(* Logix 5000 project; controller PLC_MCC1201_220AP1 vendor 1 type 14 code 164 rev 35.11; software revision 35.00; part 7 of 25 *)
(* tags used below, declared in another part *)
   B3 : DINT[102];
   HMI_Alarm_Reset : BOOL;   // HMI_Alarm_Reset
   HMI_MAN_CMD_WR : UDT_MAN_CMD_WR;
   LEHR_SPEED : ALIAS FOR N60[1];
   M210_M1_DR : AXIS_CIP_DRIVE;
   M211_M1_DR : AXIS_CIP_DRIVE;
   M212_M1_DR : AXIS_CIP_DRIVE;
   M213_M1_DR : AXIS_CIP_DRIVE;
   M2xx_CONVEYOR : MAC_CONVEYOR[20];
   M2xx_CONVEYOR_IN_MOTION : MAC_CONVEYOR_IN_MOTION[20];
   M2xx_CONVEYOR_OUT_MOTION : MAC_CONVEYOR_OUT_MOTION[20];
   TMP_dDirection : DINT;
   TMP_rAcc : REAL;
   TMP_rDec : REAL;
   TMP_rSpeed : REAL;
   TMP_xAlwaysOFF : BOOL;
   TMP_xRun : BOOL;
(* CommandLogic, continued *)

ROUTINE M210_Conveyor_Motion_Output   (* ladder *)
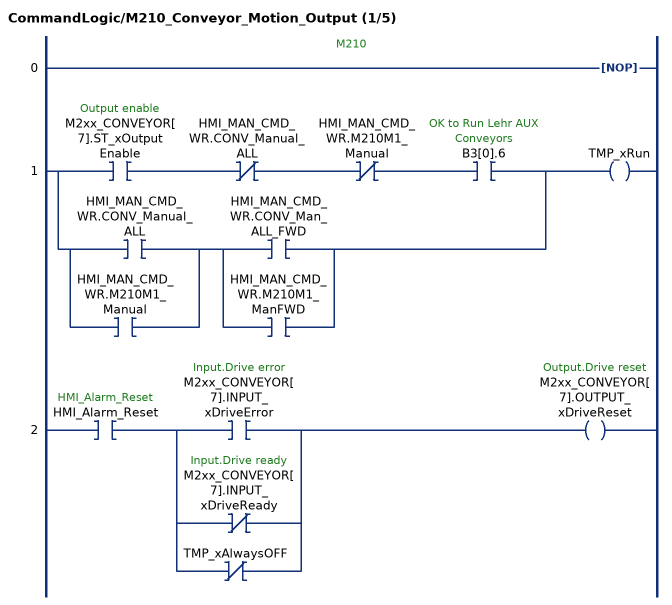
   // M210
   0: NOP();
   1: [XIC(M2xx_CONVEYOR[7].ST_xOutputEnable) XIO(HMI_MAN_CMD_WR.CONV_Manual_ALL) XIO(HMI_MAN_CMD_WR.M210M1_Manual) XIC(B3[0].6) ,[XIC(HMI_MAN_CMD_WR.CONV_Manual_ALL) ,XIC(HMI_MAN_CMD_WR.M210M1_Manual) ] [XIC(HMI_MAN_CMD_WR.CONV_Man_ALL_FWD) ,XIC(HMI_MAN_CMD_WR.M210M1_ManFWD) ] ]OTE(TMP_xRun);
   2: XIC(HMI_Alarm_Reset)[XIC(M2xx_CONVEYOR[7].INPUT_xDriveError) ,XIO(M2xx_CONVEYOR[7].INPUT_xDriveReady) ,XIO(TMP_xAlwaysOFF) ]OTE(M2xx_CONVEYOR[7].OUTPUT_xDriveReset);
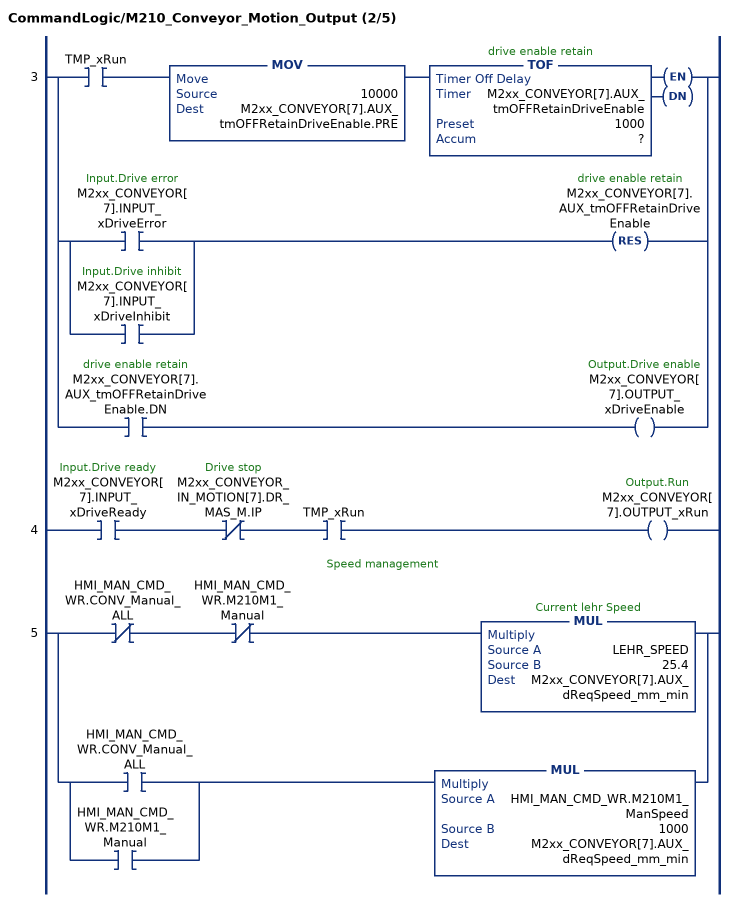
   3: [XIC(TMP_xRun) MOV(10000,M2xx_CONVEYOR[7].AUX_tmOFFRetainDriveEnable.PRE) TOF(M2xx_CONVEYOR[7].AUX_tmOFFRetainDriveEnable,?,?) ,[XIC(M2xx_CONVEYOR[7].INPUT_xDriveError) ,XIC(M2xx_CONVEYOR[7].INPUT_xDriveInhibit) ] RES(M2xx_CONVEYOR[7].AUX_tmOFFRetainDriveEnable) ,XIC(M2xx_CONVEYOR[7].AUX_tmOFFRetainDriveEnable.DN) OTE(M2xx_CONVEYOR[7].OUTPUT_xDriveEnable) ];
   4: XIC(M2xx_CONVEYOR[7].INPUT_xDriveReady)XIO(M2xx_CONVEYOR_IN_MOTION[7].DR_MAS_M.IP)XIC(TMP_xRun)OTE(M2xx_CONVEYOR[7].OUTPUT_xRun);
   // Speed management
   5: [XIO(HMI_MAN_CMD_WR.CONV_Manual_ALL) XIO(HMI_MAN_CMD_WR.M210M1_Manual) MUL(LEHR_SPEED,25.4,M2xx_CONVEYOR[7].AUX_dReqSpeed_mm_min) ,[XIC(HMI_MAN_CMD_WR.CONV_Manual_ALL) ,XIC(HMI_MAN_CMD_WR.M210M1_Manual) ] MUL(HMI_MAN_CMD_WR.M210M1_ManSpeed,1000,M2xx_CONVEYOR[7].AUX_dReqSpeed_mm_min) ];
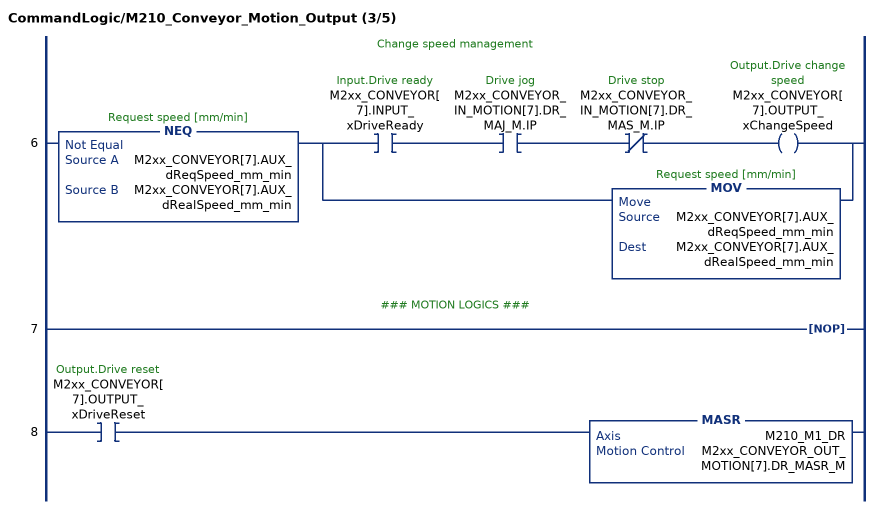
   // Change speed management
   6: NEQ(M2xx_CONVEYOR[7].AUX_dReqSpeed_mm_min,M2xx_CONVEYOR[7].AUX_dRealSpeed_mm_min)[XIC(M2xx_CONVEYOR[7].INPUT_xDriveReady) XIC(M2xx_CONVEYOR_IN_MOTION[7].DR_MAJ_M.IP) XIO(M2xx_CONVEYOR_IN_MOTION[7].DR_MAS_M.IP) OTE(M2xx_CONVEYOR[7].OUTPUT_xChangeSpeed) ,MOV(M2xx_CONVEYOR[7].AUX_dReqSpeed_mm_min,M2xx_CONVEYOR[7].AUX_dRealSpeed_mm_min) ];
   // ### MOTION LOGICS ###
   7: NOP();
   8: XIC(M2xx_CONVEYOR[7].OUTPUT_xDriveReset)MASR(M210_M1_DR,M2xx_CONVEYOR_OUT_MOTION[7].DR_MASR_M);
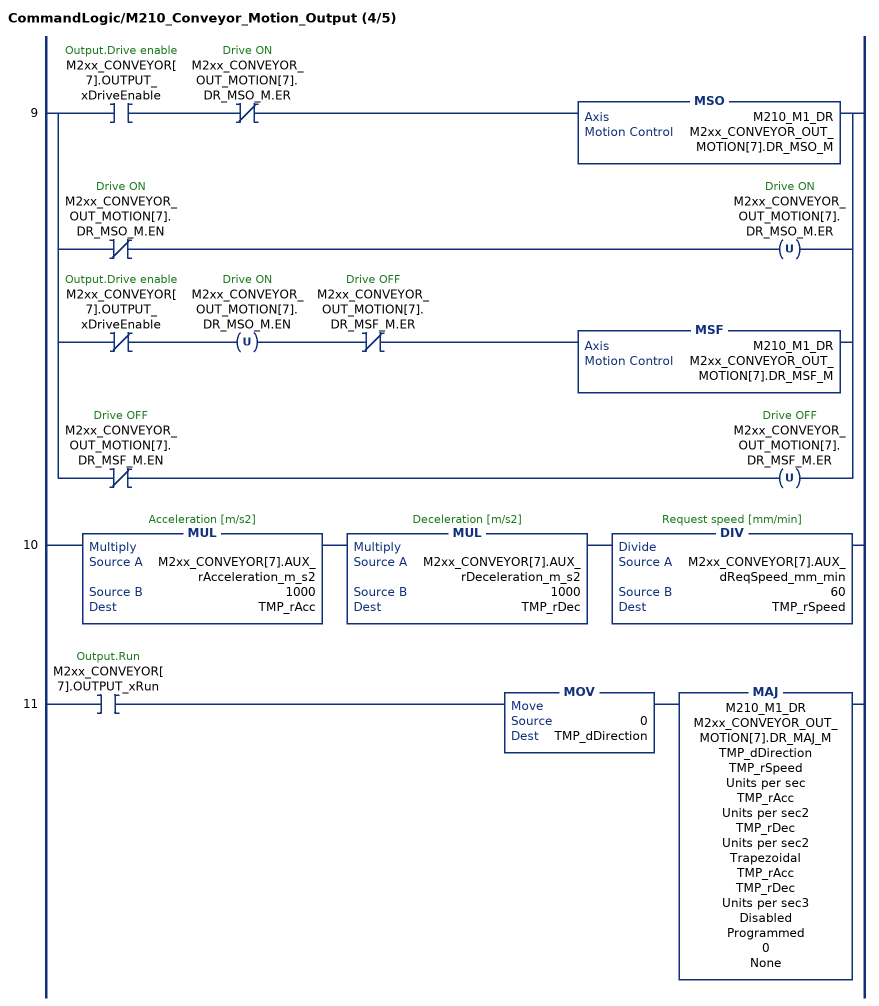
   9: [XIC(M2xx_CONVEYOR[7].OUTPUT_xDriveEnable) XIO(M2xx_CONVEYOR_OUT_MOTION[7].DR_MSO_M.ER) MSO(M210_M1_DR,M2xx_CONVEYOR_OUT_MOTION[7].DR_MSO_M) ,XIO(M2xx_CONVEYOR_OUT_MOTION[7].DR_MSO_M.EN) OTU(M2xx_CONVEYOR_OUT_MOTION[7].DR_MSO_M.ER) ,XIO(M2xx_CONVEYOR[7].OUTPUT_xDriveEnable) OTU(M2xx_CONVEYOR_OUT_MOTION[7].DR_MSO_M.EN) XIO(M2xx_CONVEYOR_OUT_MOTION[7].DR_MSF_M.ER) MSF(M210_M1_DR,M2xx_CONVEYOR_OUT_MOTION[7].DR_MSF_M) ,XIO(M2xx_CONVEYOR_OUT_MOTION[7].DR_MSF_M.EN) OTU(M2xx_CONVEYOR_OUT_MOTION[7].DR_MSF_M.ER) ];
   10: MUL(M2xx_CONVEYOR[7].AUX_rAcceleration_m_s2,1000,TMP_rAcc)MUL(M2xx_CONVEYOR[7].AUX_rDeceleration_m_s2,1000,TMP_rDec)DIV(M2xx_CONVEYOR[7].AUX_dReqSpeed_mm_min,60,TMP_rSpeed);
   11: XIC(M2xx_CONVEYOR[7].OUTPUT_xRun)MOV(0,TMP_dDirection)MAJ(M210_M1_DR,M2xx_CONVEYOR_OUT_MOTION[7].DR_MAJ_M,TMP_dDirection,TMP_rSpeed,Units per sec,TMP_rAcc,Units per sec2,TMP_rDec,Units per sec2,Trapezoidal,TMP_rAcc,TMP_rDec,Units per sec3,Disabled,Programmed,0,None);
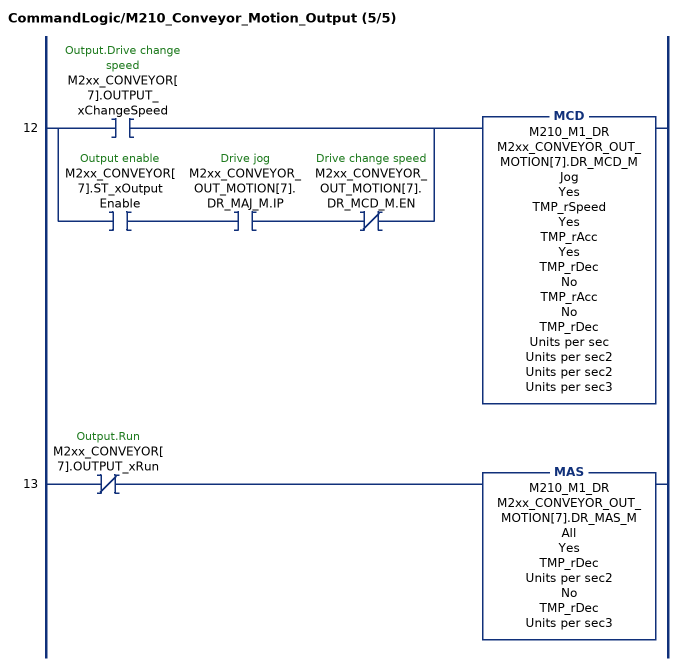
   12: [XIC(M2xx_CONVEYOR[7].OUTPUT_xChangeSpeed) ,XIC(M2xx_CONVEYOR[7].ST_xOutputEnable) XIC(M2xx_CONVEYOR_OUT_MOTION[7].DR_MAJ_M.IP) XIO(M2xx_CONVEYOR_OUT_MOTION[7].DR_MCD_M.EN) ]MCD(M210_M1_DR,M2xx_CONVEYOR_OUT_MOTION[7].DR_MCD_M,Jog,Yes,TMP_rSpeed,Yes,TMP_rAcc,Yes,TMP_rDec,No,TMP_rAcc,No,TMP_rDec,Units per sec,Units per sec2,Units per sec2,Units per sec3);
   13: XIO(M2xx_CONVEYOR[7].OUTPUT_xRun)MAS(M210_M1_DR,M2xx_CONVEYOR_OUT_MOTION[7].DR_MAS_M,All,Yes,TMP_rDec,Units per sec2,No,TMP_rDec,Units per sec3);
END_ROUTINE

ROUTINE M211_Conveyor_Motion_Output   (* ladder *)
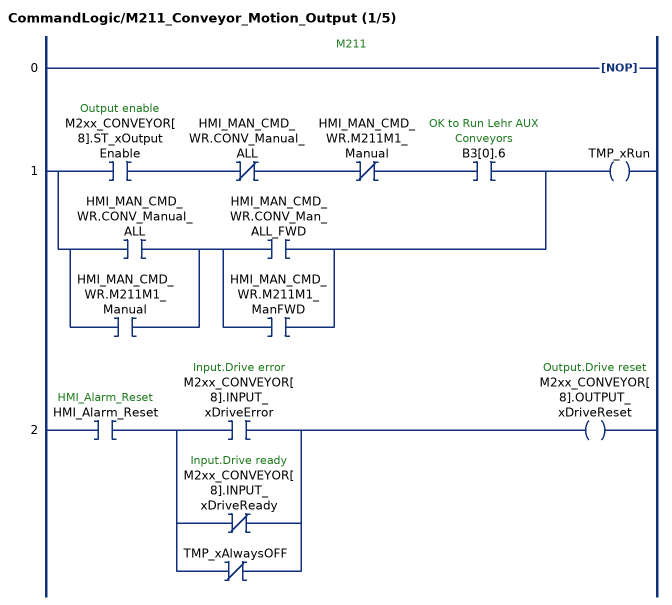
   // M211
   0: NOP();
   1: [XIC(M2xx_CONVEYOR[8].ST_xOutputEnable) XIO(HMI_MAN_CMD_WR.CONV_Manual_ALL) XIO(HMI_MAN_CMD_WR.M211M1_Manual) XIC(B3[0].6) ,[XIC(HMI_MAN_CMD_WR.CONV_Manual_ALL) ,XIC(HMI_MAN_CMD_WR.M211M1_Manual) ] [XIC(HMI_MAN_CMD_WR.CONV_Man_ALL_FWD) ,XIC(HMI_MAN_CMD_WR.M211M1_ManFWD) ] ]OTE(TMP_xRun);
   2: XIC(HMI_Alarm_Reset)[XIC(M2xx_CONVEYOR[8].INPUT_xDriveError) ,XIO(M2xx_CONVEYOR[8].INPUT_xDriveReady) ,XIO(TMP_xAlwaysOFF) ]OTE(M2xx_CONVEYOR[8].OUTPUT_xDriveReset);
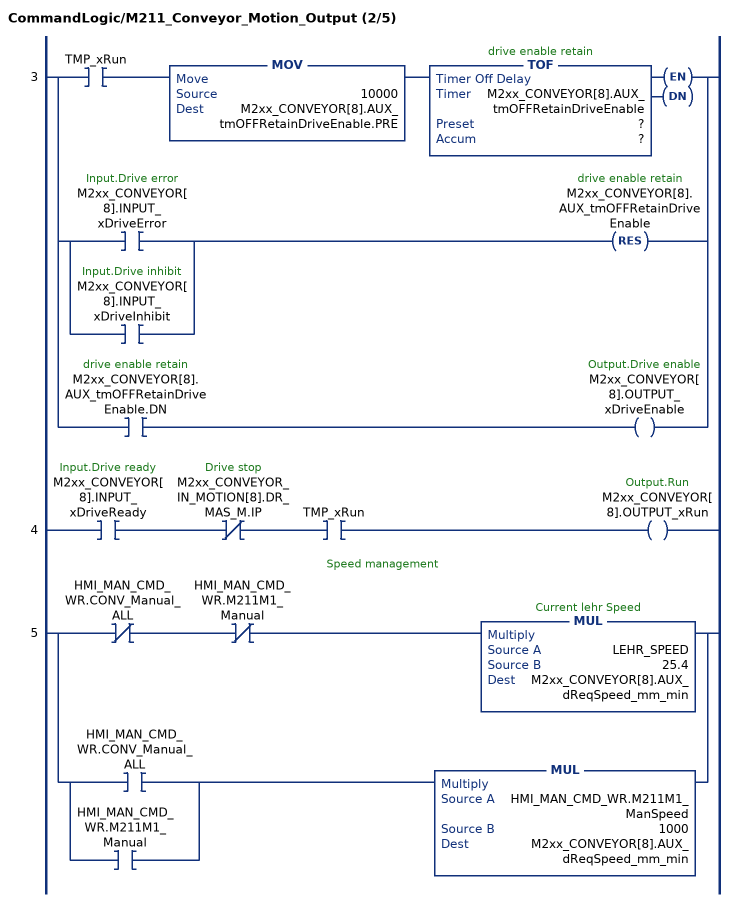
   3: [XIC(TMP_xRun) MOV(10000,M2xx_CONVEYOR[8].AUX_tmOFFRetainDriveEnable.PRE) TOF(M2xx_CONVEYOR[8].AUX_tmOFFRetainDriveEnable,?,?) ,[XIC(M2xx_CONVEYOR[8].INPUT_xDriveError) ,XIC(M2xx_CONVEYOR[8].INPUT_xDriveInhibit) ] RES(M2xx_CONVEYOR[8].AUX_tmOFFRetainDriveEnable) ,XIC(M2xx_CONVEYOR[8].AUX_tmOFFRetainDriveEnable.DN) OTE(M2xx_CONVEYOR[8].OUTPUT_xDriveEnable) ];
   4: XIC(M2xx_CONVEYOR[8].INPUT_xDriveReady)XIO(M2xx_CONVEYOR_IN_MOTION[8].DR_MAS_M.IP)XIC(TMP_xRun)OTE(M2xx_CONVEYOR[8].OUTPUT_xRun);
   // Speed management
   5: [XIO(HMI_MAN_CMD_WR.CONV_Manual_ALL) XIO(HMI_MAN_CMD_WR.M211M1_Manual) MUL(LEHR_SPEED,25.4,M2xx_CONVEYOR[8].AUX_dReqSpeed_mm_min) ,[XIC(HMI_MAN_CMD_WR.CONV_Manual_ALL) ,XIC(HMI_MAN_CMD_WR.M211M1_Manual) ] MUL(HMI_MAN_CMD_WR.M211M1_ManSpeed,1000,M2xx_CONVEYOR[8].AUX_dReqSpeed_mm_min) ];
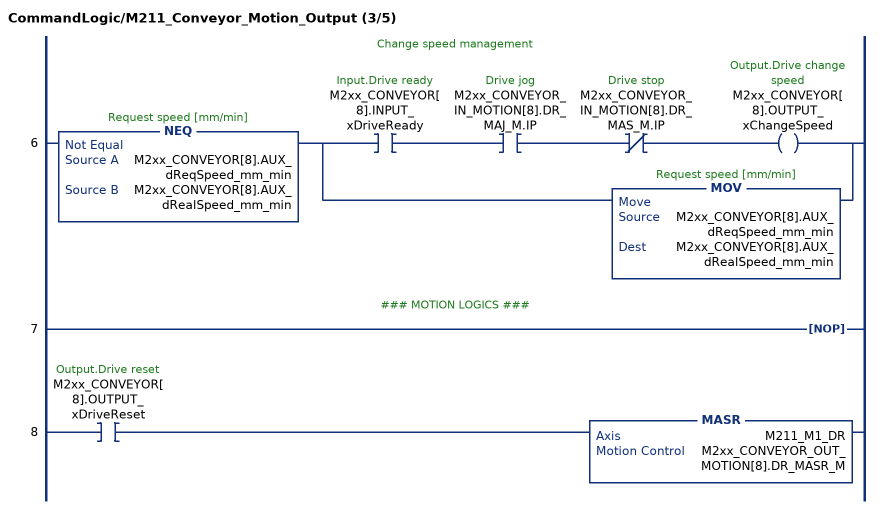
   // Change speed management
   6: NEQ(M2xx_CONVEYOR[8].AUX_dReqSpeed_mm_min,M2xx_CONVEYOR[8].AUX_dRealSpeed_mm_min)[XIC(M2xx_CONVEYOR[8].INPUT_xDriveReady) XIC(M2xx_CONVEYOR_IN_MOTION[8].DR_MAJ_M.IP) XIO(M2xx_CONVEYOR_IN_MOTION[8].DR_MAS_M.IP) OTE(M2xx_CONVEYOR[8].OUTPUT_xChangeSpeed) ,MOV(M2xx_CONVEYOR[8].AUX_dReqSpeed_mm_min,M2xx_CONVEYOR[8].AUX_dRealSpeed_mm_min) ];
   // ### MOTION LOGICS ###
   7: NOP();
   8: XIC(M2xx_CONVEYOR[8].OUTPUT_xDriveReset)MASR(M211_M1_DR,M2xx_CONVEYOR_OUT_MOTION[8].DR_MASR_M);
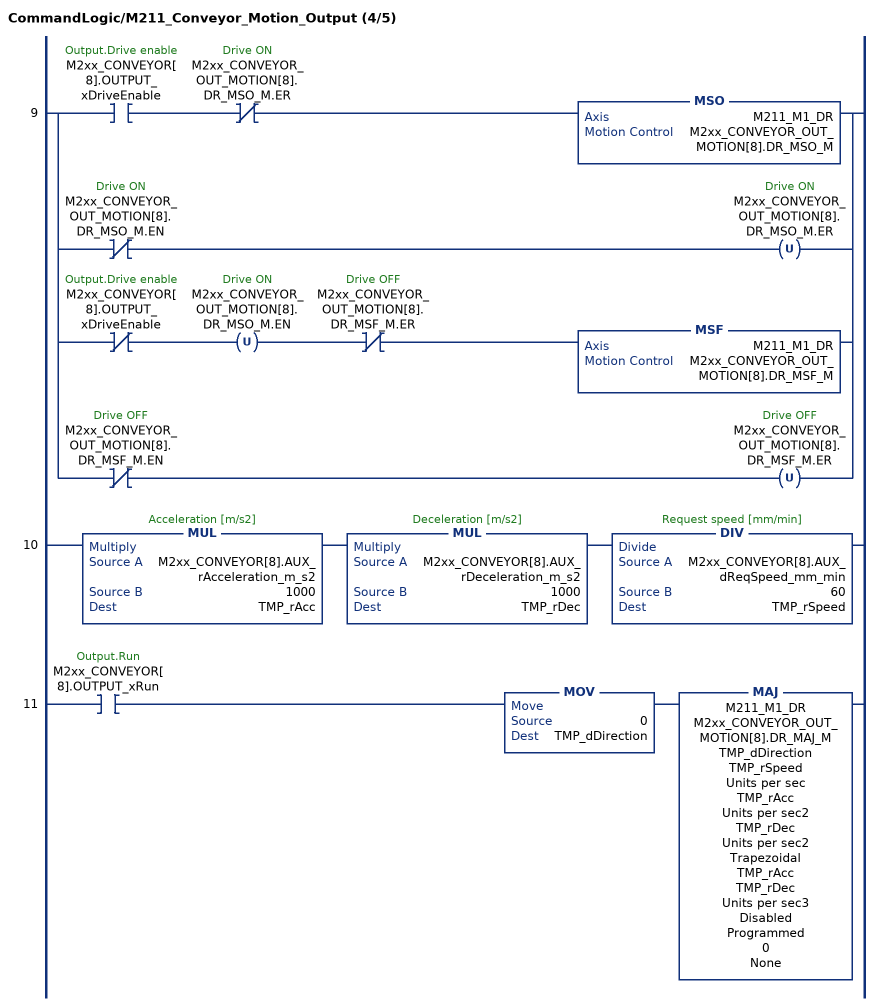
   9: [XIC(M2xx_CONVEYOR[8].OUTPUT_xDriveEnable) XIO(M2xx_CONVEYOR_OUT_MOTION[8].DR_MSO_M.ER) MSO(M211_M1_DR,M2xx_CONVEYOR_OUT_MOTION[8].DR_MSO_M) ,XIO(M2xx_CONVEYOR_OUT_MOTION[8].DR_MSO_M.EN) OTU(M2xx_CONVEYOR_OUT_MOTION[8].DR_MSO_M.ER) ,XIO(M2xx_CONVEYOR[8].OUTPUT_xDriveEnable) OTU(M2xx_CONVEYOR_OUT_MOTION[8].DR_MSO_M.EN) XIO(M2xx_CONVEYOR_OUT_MOTION[8].DR_MSF_M.ER) MSF(M211_M1_DR,M2xx_CONVEYOR_OUT_MOTION[8].DR_MSF_M) ,XIO(M2xx_CONVEYOR_OUT_MOTION[8].DR_MSF_M.EN) OTU(M2xx_CONVEYOR_OUT_MOTION[8].DR_MSF_M.ER) ];
   10: MUL(M2xx_CONVEYOR[8].AUX_rAcceleration_m_s2,1000,TMP_rAcc)MUL(M2xx_CONVEYOR[8].AUX_rDeceleration_m_s2,1000,TMP_rDec)DIV(M2xx_CONVEYOR[8].AUX_dReqSpeed_mm_min,60,TMP_rSpeed);
   11: XIC(M2xx_CONVEYOR[8].OUTPUT_xRun)MOV(0,TMP_dDirection)MAJ(M211_M1_DR,M2xx_CONVEYOR_OUT_MOTION[8].DR_MAJ_M,TMP_dDirection,TMP_rSpeed,Units per sec,TMP_rAcc,Units per sec2,TMP_rDec,Units per sec2,Trapezoidal,TMP_rAcc,TMP_rDec,Units per sec3,Disabled,Programmed,0,None);
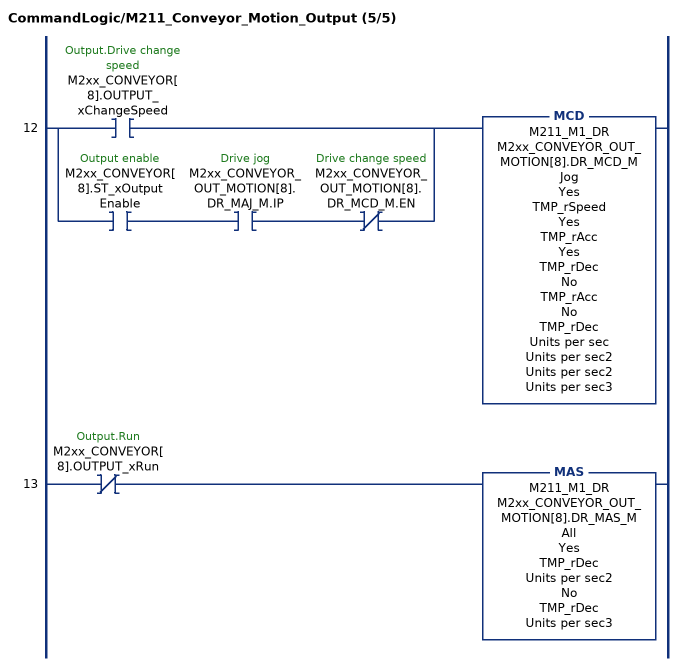
   12: [XIC(M2xx_CONVEYOR[8].OUTPUT_xChangeSpeed) ,XIC(M2xx_CONVEYOR[8].ST_xOutputEnable) XIC(M2xx_CONVEYOR_OUT_MOTION[8].DR_MAJ_M.IP) XIO(M2xx_CONVEYOR_OUT_MOTION[8].DR_MCD_M.EN) ]MCD(M211_M1_DR,M2xx_CONVEYOR_OUT_MOTION[8].DR_MCD_M,Jog,Yes,TMP_rSpeed,Yes,TMP_rAcc,Yes,TMP_rDec,No,TMP_rAcc,No,TMP_rDec,Units per sec,Units per sec2,Units per sec2,Units per sec3);
   13: XIO(M2xx_CONVEYOR[8].OUTPUT_xRun)MAS(M211_M1_DR,M2xx_CONVEYOR_OUT_MOTION[8].DR_MAS_M,All,Yes,TMP_rDec,Units per sec2,No,TMP_rDec,Units per sec3);
END_ROUTINE

ROUTINE M212_Conveyor_Motion_Output   (* ladder *)
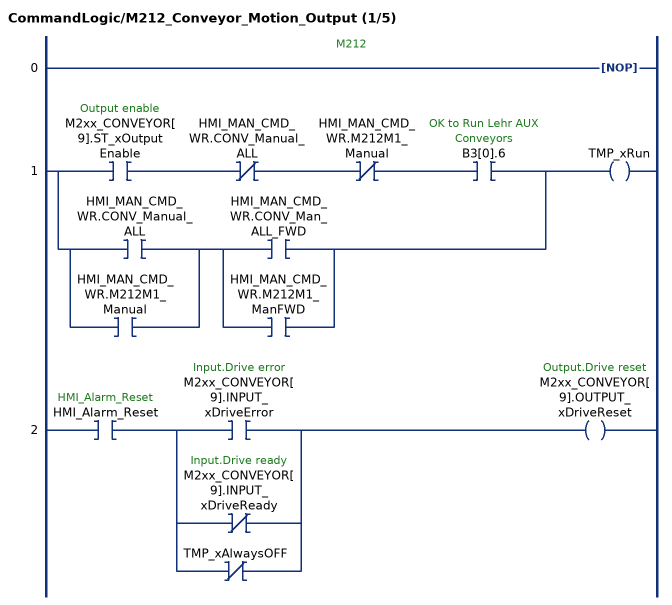
   // M212
   0: NOP();
   1: [XIC(M2xx_CONVEYOR[9].ST_xOutputEnable) XIO(HMI_MAN_CMD_WR.CONV_Manual_ALL) XIO(HMI_MAN_CMD_WR.M212M1_Manual) XIC(B3[0].6) ,[XIC(HMI_MAN_CMD_WR.CONV_Manual_ALL) ,XIC(HMI_MAN_CMD_WR.M212M1_Manual) ] [XIC(HMI_MAN_CMD_WR.CONV_Man_ALL_FWD) ,XIC(HMI_MAN_CMD_WR.M212M1_ManFWD) ] ]OTE(TMP_xRun);
   2: XIC(HMI_Alarm_Reset)[XIC(M2xx_CONVEYOR[9].INPUT_xDriveError) ,XIO(M2xx_CONVEYOR[9].INPUT_xDriveReady) ,XIO(TMP_xAlwaysOFF) ]OTE(M2xx_CONVEYOR[9].OUTPUT_xDriveReset);
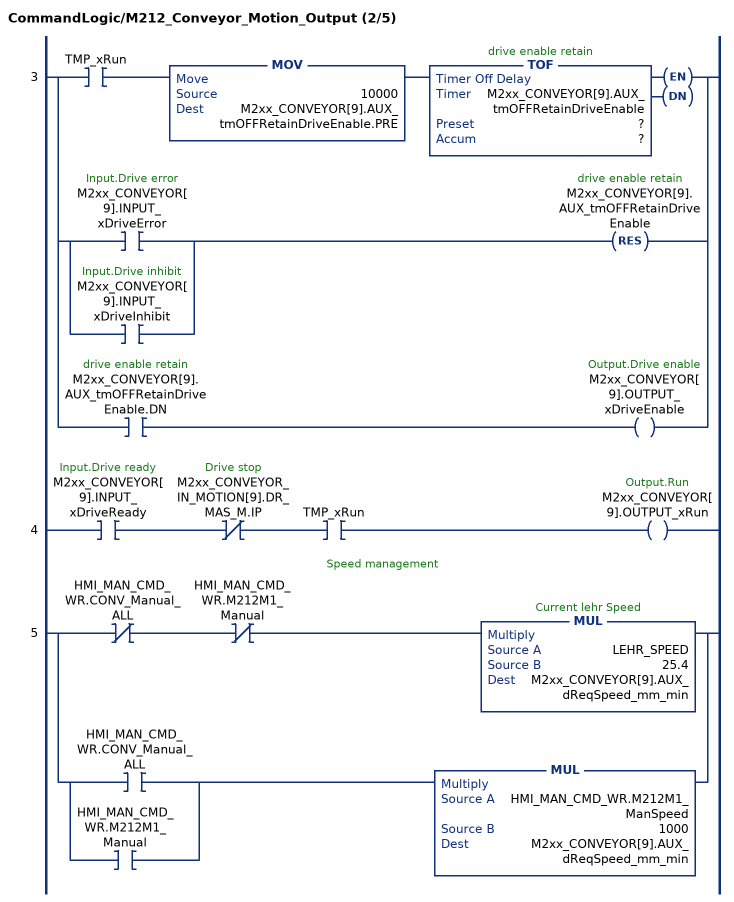
   3: [XIC(TMP_xRun) MOV(10000,M2xx_CONVEYOR[9].AUX_tmOFFRetainDriveEnable.PRE) TOF(M2xx_CONVEYOR[9].AUX_tmOFFRetainDriveEnable,?,?) ,[XIC(M2xx_CONVEYOR[9].INPUT_xDriveError) ,XIC(M2xx_CONVEYOR[9].INPUT_xDriveInhibit) ] RES(M2xx_CONVEYOR[9].AUX_tmOFFRetainDriveEnable) ,XIC(M2xx_CONVEYOR[9].AUX_tmOFFRetainDriveEnable.DN) OTE(M2xx_CONVEYOR[9].OUTPUT_xDriveEnable) ];
   4: XIC(M2xx_CONVEYOR[9].INPUT_xDriveReady)XIO(M2xx_CONVEYOR_IN_MOTION[9].DR_MAS_M.IP)XIC(TMP_xRun)OTE(M2xx_CONVEYOR[9].OUTPUT_xRun);
   // Speed management
   5: [XIO(HMI_MAN_CMD_WR.CONV_Manual_ALL) XIO(HMI_MAN_CMD_WR.M212M1_Manual) MUL(LEHR_SPEED,25.4,M2xx_CONVEYOR[9].AUX_dReqSpeed_mm_min) ,[XIC(HMI_MAN_CMD_WR.CONV_Manual_ALL) ,XIC(HMI_MAN_CMD_WR.M212M1_Manual) ] MUL(HMI_MAN_CMD_WR.M212M1_ManSpeed,1000,M2xx_CONVEYOR[9].AUX_dReqSpeed_mm_min) ];
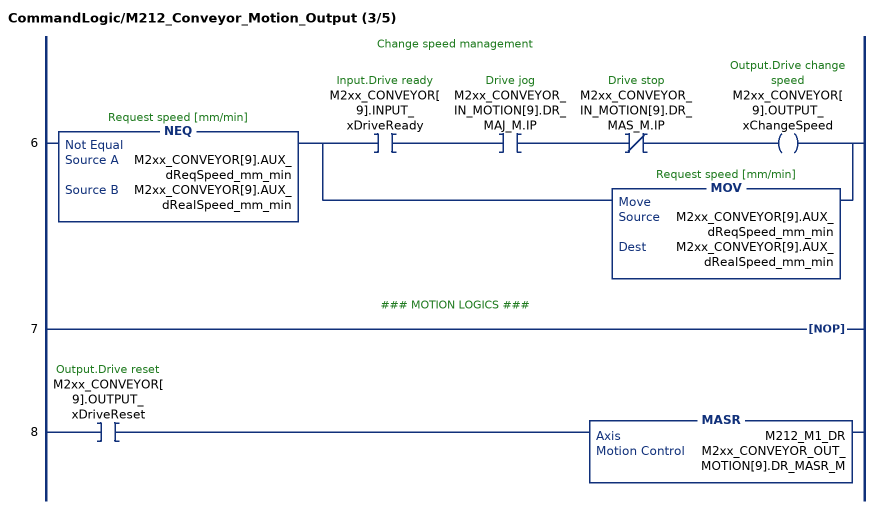
   // Change speed management
   6: NEQ(M2xx_CONVEYOR[9].AUX_dReqSpeed_mm_min,M2xx_CONVEYOR[9].AUX_dRealSpeed_mm_min)[XIC(M2xx_CONVEYOR[9].INPUT_xDriveReady) XIC(M2xx_CONVEYOR_IN_MOTION[9].DR_MAJ_M.IP) XIO(M2xx_CONVEYOR_IN_MOTION[9].DR_MAS_M.IP) OTE(M2xx_CONVEYOR[9].OUTPUT_xChangeSpeed) ,MOV(M2xx_CONVEYOR[9].AUX_dReqSpeed_mm_min,M2xx_CONVEYOR[9].AUX_dRealSpeed_mm_min) ];
   // ### MOTION LOGICS ###
   7: NOP();
   8: XIC(M2xx_CONVEYOR[9].OUTPUT_xDriveReset)MASR(M212_M1_DR,M2xx_CONVEYOR_OUT_MOTION[9].DR_MASR_M);
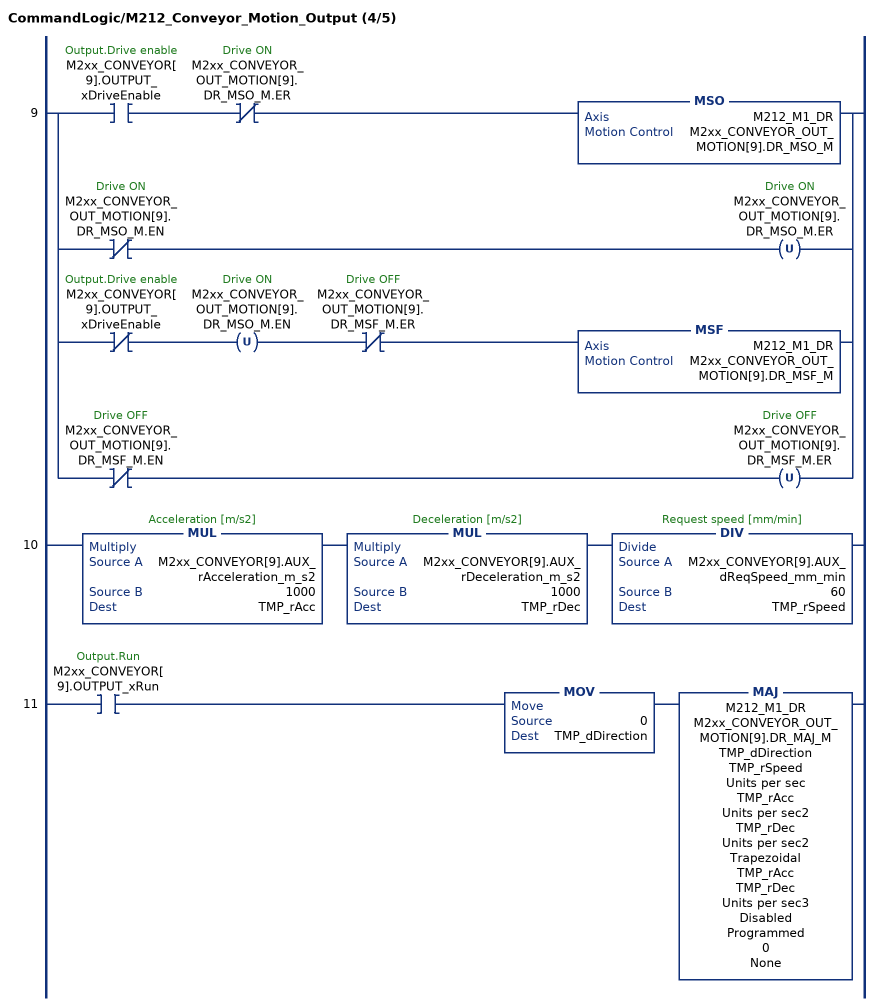
   9: [XIC(M2xx_CONVEYOR[9].OUTPUT_xDriveEnable) XIO(M2xx_CONVEYOR_OUT_MOTION[9].DR_MSO_M.ER) MSO(M212_M1_DR,M2xx_CONVEYOR_OUT_MOTION[9].DR_MSO_M) ,XIO(M2xx_CONVEYOR_OUT_MOTION[9].DR_MSO_M.EN) OTU(M2xx_CONVEYOR_OUT_MOTION[9].DR_MSO_M.ER) ,XIO(M2xx_CONVEYOR[9].OUTPUT_xDriveEnable) OTU(M2xx_CONVEYOR_OUT_MOTION[9].DR_MSO_M.EN) XIO(M2xx_CONVEYOR_OUT_MOTION[9].DR_MSF_M.ER) MSF(M212_M1_DR,M2xx_CONVEYOR_OUT_MOTION[9].DR_MSF_M) ,XIO(M2xx_CONVEYOR_OUT_MOTION[9].DR_MSF_M.EN) OTU(M2xx_CONVEYOR_OUT_MOTION[9].DR_MSF_M.ER) ];
   10: MUL(M2xx_CONVEYOR[9].AUX_rAcceleration_m_s2,1000,TMP_rAcc)MUL(M2xx_CONVEYOR[9].AUX_rDeceleration_m_s2,1000,TMP_rDec)DIV(M2xx_CONVEYOR[9].AUX_dReqSpeed_mm_min,60,TMP_rSpeed);
   11: XIC(M2xx_CONVEYOR[9].OUTPUT_xRun)MOV(0,TMP_dDirection)MAJ(M212_M1_DR,M2xx_CONVEYOR_OUT_MOTION[9].DR_MAJ_M,TMP_dDirection,TMP_rSpeed,Units per sec,TMP_rAcc,Units per sec2,TMP_rDec,Units per sec2,Trapezoidal,TMP_rAcc,TMP_rDec,Units per sec3,Disabled,Programmed,0,None);
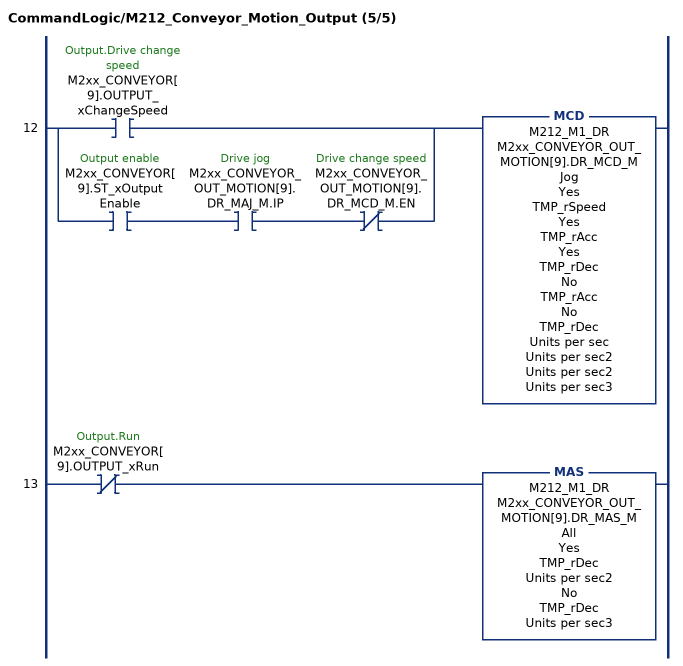
   12: [XIC(M2xx_CONVEYOR[9].OUTPUT_xChangeSpeed) ,XIC(M2xx_CONVEYOR[9].ST_xOutputEnable) XIC(M2xx_CONVEYOR_OUT_MOTION[9].DR_MAJ_M.IP) XIO(M2xx_CONVEYOR_OUT_MOTION[9].DR_MCD_M.EN) ]MCD(M212_M1_DR,M2xx_CONVEYOR_OUT_MOTION[9].DR_MCD_M,Jog,Yes,TMP_rSpeed,Yes,TMP_rAcc,Yes,TMP_rDec,No,TMP_rAcc,No,TMP_rDec,Units per sec,Units per sec2,Units per sec2,Units per sec3);
   13: XIO(M2xx_CONVEYOR[9].OUTPUT_xRun)MAS(M212_M1_DR,M2xx_CONVEYOR_OUT_MOTION[9].DR_MAS_M,All,Yes,TMP_rDec,Units per sec2,No,TMP_rDec,Units per sec3);
END_ROUTINE

ROUTINE M213_Conveyor_Motion_Output   (* ladder *)
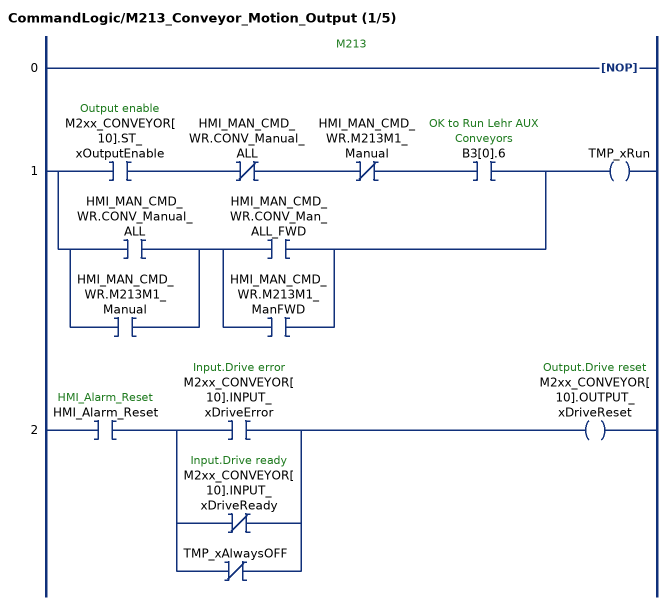
   // M213
   0: NOP();
   1: [XIC(M2xx_CONVEYOR[10].ST_xOutputEnable) XIO(HMI_MAN_CMD_WR.CONV_Manual_ALL) XIO(HMI_MAN_CMD_WR.M213M1_Manual) XIC(B3[0].6) ,[XIC(HMI_MAN_CMD_WR.CONV_Manual_ALL) ,XIC(HMI_MAN_CMD_WR.M213M1_Manual) ] [XIC(HMI_MAN_CMD_WR.CONV_Man_ALL_FWD) ,XIC(HMI_MAN_CMD_WR.M213M1_ManFWD) ] ]OTE(TMP_xRun);
   2: XIC(HMI_Alarm_Reset)[XIC(M2xx_CONVEYOR[10].INPUT_xDriveError) ,XIO(M2xx_CONVEYOR[10].INPUT_xDriveReady) ,XIO(TMP_xAlwaysOFF) ]OTE(M2xx_CONVEYOR[10].OUTPUT_xDriveReset);
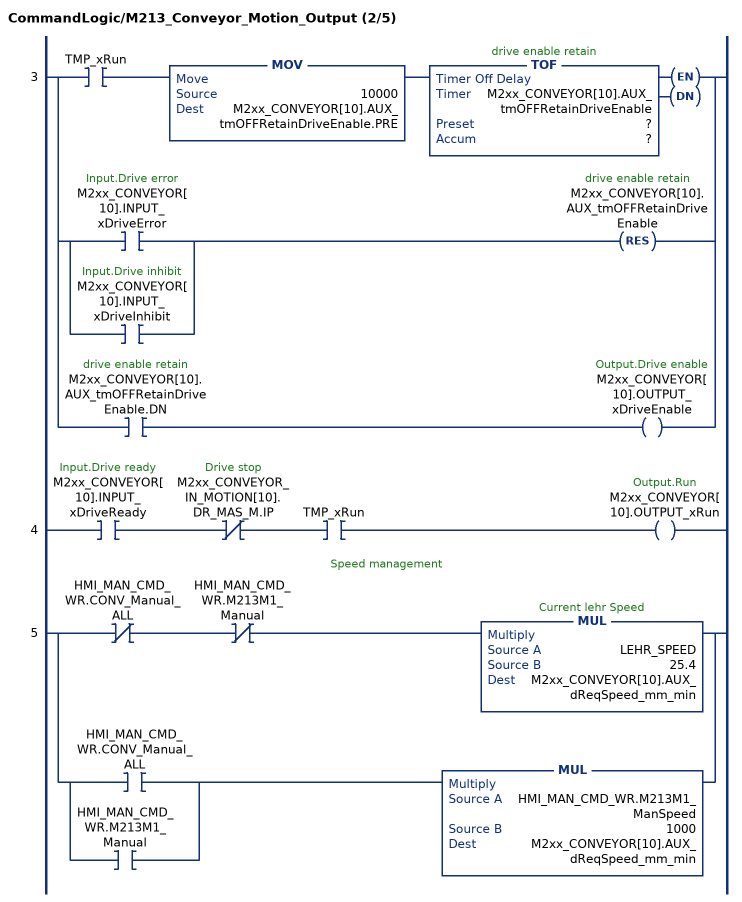
   3: [XIC(TMP_xRun) MOV(10000,M2xx_CONVEYOR[10].AUX_tmOFFRetainDriveEnable.PRE) TOF(M2xx_CONVEYOR[10].AUX_tmOFFRetainDriveEnable,?,?) ,[XIC(M2xx_CONVEYOR[10].INPUT_xDriveError) ,XIC(M2xx_CONVEYOR[10].INPUT_xDriveInhibit) ] RES(M2xx_CONVEYOR[10].AUX_tmOFFRetainDriveEnable) ,XIC(M2xx_CONVEYOR[10].AUX_tmOFFRetainDriveEnable.DN) OTE(M2xx_CONVEYOR[10].OUTPUT_xDriveEnable) ];
   4: XIC(M2xx_CONVEYOR[10].INPUT_xDriveReady)XIO(M2xx_CONVEYOR_IN_MOTION[10].DR_MAS_M.IP)XIC(TMP_xRun)OTE(M2xx_CONVEYOR[10].OUTPUT_xRun);
   // Speed management
   5: [XIO(HMI_MAN_CMD_WR.CONV_Manual_ALL) XIO(HMI_MAN_CMD_WR.M213M1_Manual) MUL(LEHR_SPEED,25.4,M2xx_CONVEYOR[10].AUX_dReqSpeed_mm_min) ,[XIC(HMI_MAN_CMD_WR.CONV_Manual_ALL) ,XIC(HMI_MAN_CMD_WR.M213M1_Manual) ] MUL(HMI_MAN_CMD_WR.M213M1_ManSpeed,1000,M2xx_CONVEYOR[10].AUX_dReqSpeed_mm_min) ];
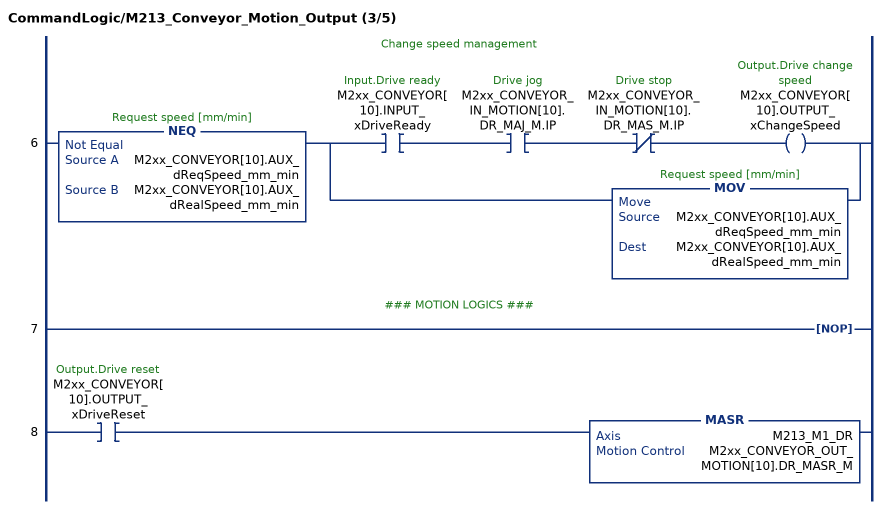
   // Change speed management
   6: NEQ(M2xx_CONVEYOR[10].AUX_dReqSpeed_mm_min,M2xx_CONVEYOR[10].AUX_dRealSpeed_mm_min)[XIC(M2xx_CONVEYOR[10].INPUT_xDriveReady) XIC(M2xx_CONVEYOR_IN_MOTION[10].DR_MAJ_M.IP) XIO(M2xx_CONVEYOR_IN_MOTION[10].DR_MAS_M.IP) OTE(M2xx_CONVEYOR[10].OUTPUT_xChangeSpeed) ,MOV(M2xx_CONVEYOR[10].AUX_dReqSpeed_mm_min,M2xx_CONVEYOR[10].AUX_dRealSpeed_mm_min) ];
   // ### MOTION LOGICS ###
   7: NOP();
   8: XIC(M2xx_CONVEYOR[10].OUTPUT_xDriveReset)MASR(M213_M1_DR,M2xx_CONVEYOR_OUT_MOTION[10].DR_MASR_M);
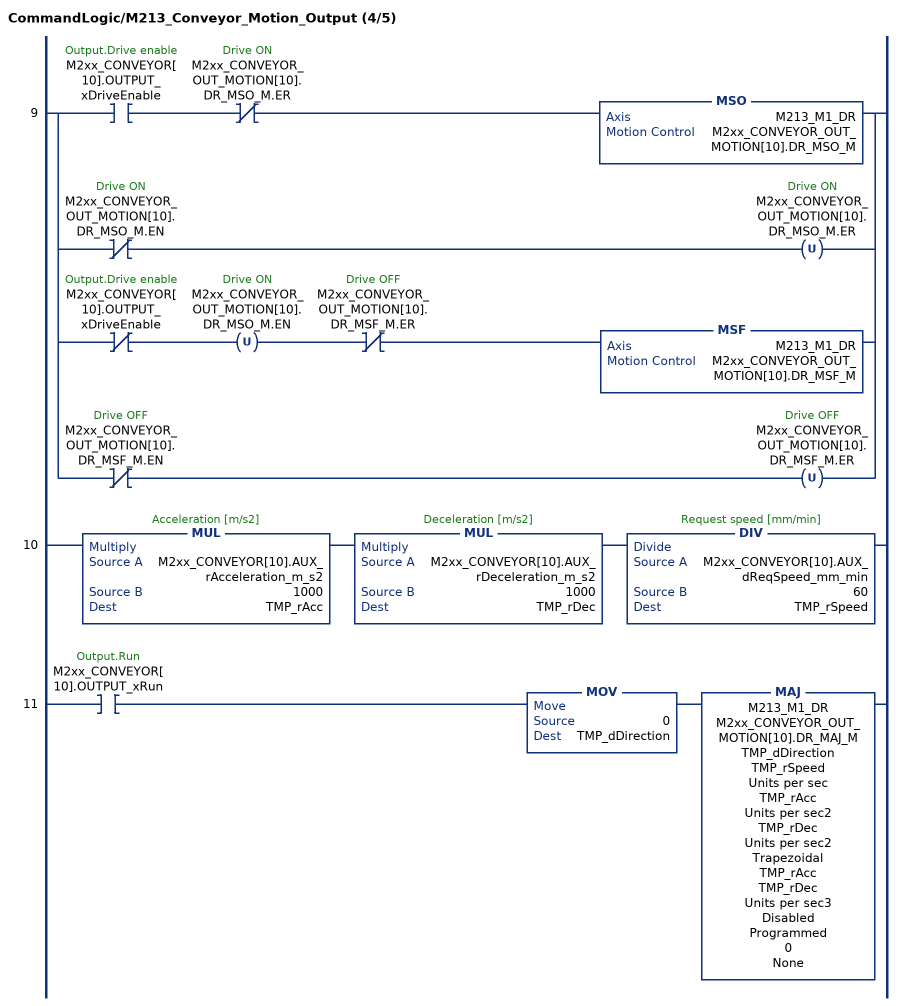
   9: [XIC(M2xx_CONVEYOR[10].OUTPUT_xDriveEnable) XIO(M2xx_CONVEYOR_OUT_MOTION[10].DR_MSO_M.ER) MSO(M213_M1_DR,M2xx_CONVEYOR_OUT_MOTION[10].DR_MSO_M) ,XIO(M2xx_CONVEYOR_OUT_MOTION[10].DR_MSO_M.EN) OTU(M2xx_CONVEYOR_OUT_MOTION[10].DR_MSO_M.ER) ,XIO(M2xx_CONVEYOR[10].OUTPUT_xDriveEnable) OTU(M2xx_CONVEYOR_OUT_MOTION[10].DR_MSO_M.EN) XIO(M2xx_CONVEYOR_OUT_MOTION[10].DR_MSF_M.ER) MSF(M213_M1_DR,M2xx_CONVEYOR_OUT_MOTION[10].DR_MSF_M) ,XIO(M2xx_CONVEYOR_OUT_MOTION[10].DR_MSF_M.EN) OTU(M2xx_CONVEYOR_OUT_MOTION[10].DR_MSF_M.ER) ];
   10: MUL(M2xx_CONVEYOR[10].AUX_rAcceleration_m_s2,1000,TMP_rAcc)MUL(M2xx_CONVEYOR[10].AUX_rDeceleration_m_s2,1000,TMP_rDec)DIV(M2xx_CONVEYOR[10].AUX_dReqSpeed_mm_min,60,TMP_rSpeed);
   11: XIC(M2xx_CONVEYOR[10].OUTPUT_xRun)MOV(0,TMP_dDirection)MAJ(M213_M1_DR,M2xx_CONVEYOR_OUT_MOTION[10].DR_MAJ_M,TMP_dDirection,TMP_rSpeed,Units per sec,TMP_rAcc,Units per sec2,TMP_rDec,Units per sec2,Trapezoidal,TMP_rAcc,TMP_rDec,Units per sec3,Disabled,Programmed,0,None);
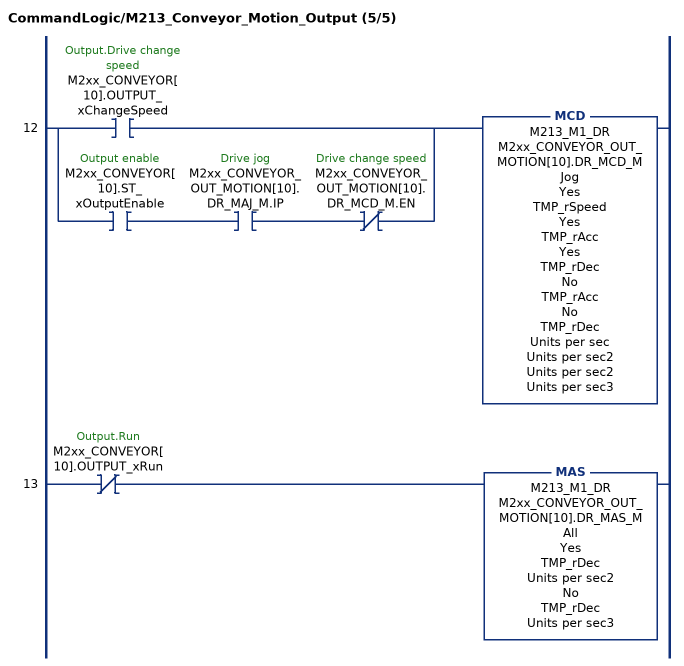
   12: [XIC(M2xx_CONVEYOR[10].OUTPUT_xChangeSpeed) ,XIC(M2xx_CONVEYOR[10].ST_xOutputEnable) XIC(M2xx_CONVEYOR_OUT_MOTION[10].DR_MAJ_M.IP) XIO(M2xx_CONVEYOR_OUT_MOTION[10].DR_MCD_M.EN) ]MCD(M213_M1_DR,M2xx_CONVEYOR_OUT_MOTION[10].DR_MCD_M,Jog,Yes,TMP_rSpeed,Yes,TMP_rAcc,Yes,TMP_rDec,No,TMP_rAcc,No,TMP_rDec,Units per sec,Units per sec2,Units per sec2,Units per sec3);
   13: XIO(M2xx_CONVEYOR[10].OUTPUT_xRun)MAS(M213_M1_DR,M2xx_CONVEYOR_OUT_MOTION[10].DR_MAS_M,All,Yes,TMP_rDec,Units per sec2,No,TMP_rDec,Units per sec3);
END_ROUTINE
